// TIA Portal project "DHARMA_1500" (V15) (continued)
VAR_GLOBAL   // PLC tag table "I/O-TurnTable"
   "TT_ES_Operatingpanel" AT %I1104.0 : Bool;   // Turntable: Emergency stop control panel
   "TT_F_CircuitBreaker" AT %I1100.0 : Bool;   // Turntable: Fault supply
   "TT_T_Start" AT %I1104.1 : Bool;   // Turntable: Start automatic
   "TT_T_Stop" AT %I1104.2 : Bool;   // Turntable: Stop automatic
   "TT_T_Reference" AT %I104.5 : Bool;   // Taster zum Turntable: Referezpunktfahren des Rundtisches "Referenzieren"
   "TT_T_TipTT+" AT %I1104.3 : Bool;   // Turntable: Taster Tippen "+" Rundtisch
   "TT_T_TipTT-" AT %I1104.4 : Bool;   // Turntable: Taster Tippen "-" Rundtisch
   "TT_S_OM_Manual" AT %I104.7 : Bool;   // Schlüsselschalter Rundtisch auf Handbetrieb
   "TT_S_OM_Auto" AT %I104.6 : Bool;   // Schlüsselschalter Rundtisch auf Automatikbetrieb
   "TT_B_Empty" AT %I1105.0 : Bool;   // Taster "Leerfahren"
   "TT_B_WithoutFoam" AT %I1105.1 : Bool;   // Taster "ohne schäumen"
   "TT_F_Supply_FC" AT %I1102.4 : Bool;   // Störung der Versorgung des Frequenzumrichters des Rundtisches
   "TT_F_FC" AT %I1101.0 : Bool;   // Turntable: Fault from frequency converter
   "TT_LS_ToolExist" AT %I1102.6 : Bool;   // Lichtschranke Werkzeug bvorhanden
   "TT_LS_ToolClose" AT %I1102.7 : Bool;   // Lichtschranke Werkzeug geschlossen
   "TT_S_SelectDoor_1" AT %I1102.3 : Bool;   // Turntable: Select open door 1
   "TT_AS_WingDoor" AT %I1100.3 : Bool;   // Turntable: Wing dooor rady
   "TT_AS" AT %I1100.7 : Bool;   // Turntable: Automatic stop ready
   "E_MK_Reiniger_Zyl_Aus" AT %I1107.0 : Bool;   // Zylinder 1 Reiniger Mischkopf ausgefahren
   "E_MK_Reiniger_Zyl_Ein" AT %I1107.1 : Bool;   // Zylinder 1 Reiniger Mischkopf eingefahren
   "T_MK_Reiniger_in_GS" AT %I1106.4 : Bool;   // Taster Mischkopfreiniger in Grundstellung fahren
   "T_MK_Reiniger_in_AS" AT %I1106.5 : Bool;   // Taster Mischkopfreiniger in Arbeitsstellung fahren
   "TT_in_position" AT %I1102.5 : Bool;   // Signal "Genauhalt" Rundtisch
   "P_MK_Reiniger_Zyl" AT %I1107.2 : Bool;   // Zylinder 1 Reiniger Mischkopf Druckluft vorhanden
   "TT_Enable_FC" AT %Q104.4 : Bool;   // Ansteuerunr des Umrichters für den Rundtisch
   "TT_V_OpenDoor_1" AT %Q104.2 : Bool;   // Turntable: Clamping valve door 1
   "TT_H_ReleaseDoor_1" AT %Q104.3 : Bool;   // Turntable: Light door 1
   "TT_H_AS" AT %Q105.7 : Bool;   // Turntable: Light automatik stop ready
   "TT_H_Start" AT %Q104.0 : Bool;   // Anzeige zum starten der Anlage
   "TT_H_Anfahrwarnung" AT %Q104.7 : Bool;
   "TT_H_Tip+" AT %Q105.4 : Bool;
   "TT_H_Tip-" AT %Q105.5 : Bool;
   "TT_H_Reference" AT %Q105.6 : Bool;
END_VAR

VAR_GLOBAL   // PLC tag table "I/O TT main"
   "F_fuse_machine(1)" AT %I100.2 : Bool;
   "F_fuse_slip_ring" AT %I100.3 : Bool;
   "ES_turn_table" AT %I100.4 : Bool;
   "AS_turn_table" AT %I100.7 : Bool;
   "F_cooling_unit" AT %I100.5 : Bool;
   "F_fuse_robot" AT %I100.6 : Bool;
   "F_FC_turn_table" AT %I107.0 : Bool;
   "F_fuse_FC_turn_table" AT %I107.1 : Bool;
   "F_fuse_24V_TT_main" AT %I100.1 : Bool;
   "ES_TT_main_cabinet" AT %I101.0 : Bool;
   "ES_TT_operating_panel" AT %I101.1 : Bool;
   "ES_TT_removal_area" AT %I101.2 : Bool;
   "ES_TT_tool_change" AT %I101.3 : Bool;
   "ES_TT_safety_door_robot" AT %I101.4 : Bool;
   "ES_TT_limit_switch_chain" AT %I101.5 : Bool;
   "Controlvoltage_okay" AT %I100.0 : Bool;
   "AS_door_tool_change" AT %I102.0 : Bool;
   "Quit_door_tool_change" AT %I102.1 : Bool;
   "Select_door_tool_change" AT %I102.2 : Bool;
   "AS_door_robot" AT %I102.3 : Bool;
   "Quit_door_robot" AT %I102.4 : Bool;
   "Select_door_robot" AT %I102.5 : Bool;
   "AS_pendelum_flap_to_handling" AT %I102.6 : Bool;
   "AS_pendelum_flap_from_handling" AT %I102.7 : Bool;
   "AS_Scanner_handling" AT %I103.0 : Bool;
   "Button_slider_HP" AT %I103.1 : Bool;
   "Button_slider_WP" AT %I103.2 : Bool;
   "Scanner_dirty" AT %I103.3 : Bool;
   "ES_robot" AT %I101.6 : Bool;
   "AS_robot_safety_area_1" AT %I103.6 : Bool;
   "AS_okay" AT %I103.7 : Bool;
   "ES_foaming_machine" AT %I101.7 : Bool;
   "I_exact_stop_TT" AT %I107.2 : Bool;
   "P_chain_tensioner" AT %I107.3 : Bool;
   "Quit_fault" AT %I104.4 : Bool;
   "Switch_manual_mode" AT %I104.0 : Bool;
   "Switch_automatic_mode" AT %I104.1 : Bool;
   "Button_start_cycle" AT %I104.2 : Bool;
   "Button_stop_cycle" AT %I104.3 : Bool;
   "Button_reference_TT" AT %I105.1 : Bool;
   "Button_TT_empty" AT %I105.2 : Bool;
   "Button_Tip_+" AT %I105.3 : Bool;
   "Button_Tip_-" AT %I105.4 : Bool;
   "Button_extend_cycle" AT %I105.5 : Bool;
   "Button_without_foam" AT %I105.0 : Bool;
   "Button_Move_+" AT %I105.6 : Bool;
   "Button_Move_-" AT %I105.7 : Bool;
   "BCD_Movement_Bit_0" AT %I106.0 : Bool;
   "BCD_Movement_Bit_1" AT %I106.1 : Bool;
   "BCD_Movement_Bit_2" AT %I106.2 : Bool;
   "BCD_Movement_Bit_3" AT %I106.3 : Bool;
   "BCD_MC_Bit_0" AT %I106.4 : Bool;
   "BCD_MC_Bit_1" AT %I106.5 : Bool;
   "BCD_MC_Bit_2" AT %I106.6 : Bool;
   "BCD_MC_Bit_3" AT %I106.7 : Bool;
   "BCD_Movement_MC" AT %IB106 : Byte;
   "Release_FC_turn_table" AT %Q103.7 : Bool;
   "Release_door_tool_change" AT %Q103.0 : Bool;
   "Selected_door_tool_change" AT %Q100.0 : Bool;
   "Release_door_robot" AT %Q103.1 : Bool;
   "Selected_door_robot" AT %Q100.1 : Bool;
   "Quit_scanner_handling" AT %Q100.7 : Bool;
   "LED_slider_HP" AT %Q102.1 : Bool;
   "LED_slider_WP" AT %Q102.2 : Bool;
   "Quit_automatic_stop" AT %Q100.2 : Bool;
   "V_chain_tensioner" AT %Q102.7 : Bool;
   "LED_start_cycle" AT %Q101.0 : Bool;
   "LED_reference_TT" AT %Q101.1 : Bool;
   "LED_TT_empty" AT %Q101.2 : Bool;
   "LED_Tip_+" AT %Q101.3 : Bool;
   "LED_Tip_-" AT %Q101.4 : Bool;
   "LED_extend_cycle" AT %Q101.5 : Bool;
   "LED_Move_+" AT %Q101.6 : Bool;
   "LED_Move_-" AT %Q101.7 : Bool;
   "Horn_TT_start" AT %Q100.3 : Bool;
   "LED_fault" AT %Q100.5 : Bool;
   "Horn_fault" AT %Q100.6 : Bool;
   "LED_TT_ready" AT %Q100.4 : Bool;
END_VAR

VAR_GLOBAL   // PLC tag table "Generell"
   "Flag_10_000_Hertz" AT %M0.0 : Bool;   // System flag of pulse 10.000 Hertz
   "Flag_05_000_Hertz" AT %M0.1 : Bool;   // System flag of pulse 5.000 Hertz
   "Flag_02_500_Hertz" AT %M0.2 : Bool;   // System flag of pulse 2.500 Hertz
   "Flag_02_000_Hertz" AT %M0.3 : Bool;   // System flag of pulse 2.000 Hertz
   "Flag_01_250_Hertz" AT %M0.4 : Bool;   // System flag of pulse 1.250 Hertz
   "Flag_01_000_Hertz" AT %M0.5 : Bool;   // System flag of pulse 1.000 Hertz
   "Flag_00_625_Hertz" AT %M0.6 : Bool;   // System flag of pulse 0.625 Hertz
   "Flag_00_500_Hertz" AT %M0.7 : Bool;   // System flag of pulse 0.500 Hertz
   "Flag_Erster_SPS_Zyklus" AT %M2.1 : Bool;   // Flag first plc cycle running
   "Flag_DP_Bus1_ADR001_ok" AT %M10.0 : Bool;   // profibus member at DP-Bus 01 with address 001 is available
   "Flag_DP_Bus1_ADR002_ok" AT %M10.1 : Bool;   // profibus member at DP-Bus 01 with address 002 is available
   "Flag_DP_Bus1_ADR003_ok" AT %M10.2 : Bool;   // profibus member at DP-Bus 01 with address 003 is available
   "Flag_DP_Bus1_ADR004_ok" AT %M10.3 : Bool;   // profibus member at DP-Bus 01 with address 004 is available
   "Flag_DP_Bus1_ADR005_ok" AT %M10.4 : Bool;   // profibus member at DP-Bus 01 with address 005 is available
   "Flag_DP_Bus1_ADR006_ok" AT %M10.5 : Bool;   // profibus member at DP-Bus 01 with address 006 is available
   "Flag_DP_Bus1_ADR007_ok" AT %M10.6 : Bool;   // profibus member at DP-Bus 01 with address 007 is available
   "Flag_DP_Bus1_ADR008_ok" AT %M10.7 : Bool;   // profibus member at DP-Bus 01 with address 008 is available
   "Flag_DP_Bus1_ADR009_ok" AT %M11.0 : Bool;   // profibus member at DP-Bus 01 with address 009 is available
   "Flag_DP_Bus1_ADR010_ok" AT %M11.1 : Bool;   // profibus member at DP-Bus 01 with address 010 is available
   "Flag_DP_Bus1_ADR011_ok" AT %M11.2 : Bool;   // profibus member at DP-Bus 01 with address 011 is available
   "Flag_DP_Bus1_ADR012_ok" AT %M11.3 : Bool;   // profibus member at DP-Bus 01 with address 012 is available
   "Flag_DP_Bus1_ADR013_ok" AT %M11.4 : Bool;   // profibus member at DP-Bus 01 with address 013 is available
   "Flag_DP_Bus1_ADR014_ok" AT %M11.5 : Bool;   // profibus member at DP-Bus 01 with address 014 is available
   "Flag_DP_Bus1_ADR015_ok" AT %M11.6 : Bool;   // profibus member at DP-Bus 01 with address 015 is available
   "Flag_DP_Bus1_ADR016_ok" AT %M11.7 : Bool;   // profibus member at DP-Bus 01 with address 016 is available
   "Flag_DP_Bus1_ADR017_ok" AT %M12.0 : Bool;   // profibus member at DP-Bus 01 with address 017 is available
   "Flag_DP_Bus1_ADR018_ok" AT %M12.1 : Bool;   // profibus member at DP-Bus 01 with address 018 is available
   "Flag_DP_Bus1_ADR019_ok" AT %M12.2 : Bool;   // profibus member at DP-Bus 01 with address 019 is available
   "Flag_DP_Bus1_ADR020_ok" AT %M12.3 : Bool;   // profibus member at DP-Bus 01 with address 020 is available
   "Flag_DP_Bus1_ADR021_ok" AT %M12.4 : Bool;   // profibus member at DP-Bus 01 with address 021 is available
   "Flag_DP_Bus1_ADR022_ok" AT %M12.5 : Bool;   // profibus member at DP-Bus 01 with address 022 is available
   "Flag_DP_Bus1_ADR023_ok" AT %M12.6 : Bool;   // profibus member at DP-Bus 01 with address 023 is available
   "Flag_DP_Bus1_ADR024_ok" AT %M12.7 : Bool;   // profibus member at DP-Bus 01 with address 024 is available
   "Flag_DP_Bus1_ADR025_ok" AT %M13.0 : Bool;   // profibus member at DP-Bus 01 with address 025 is available
   "Flag_DP_Bus1_ADR026_ok" AT %M13.1 : Bool;   // profibus member at DP-Bus 01 with address 026 is available
   "Flag_DP_Bus1_ADR027_ok" AT %M13.2 : Bool;   // profibus member at DP-Bus 01 with address 027 is available
   "Flag_DP_Bus1_ADR028_ok" AT %M13.3 : Bool;   // profibus member at DP-Bus 01 with address 028 is available
   "Flag_DP_Bus1_ADR029_ok" AT %M13.4 : Bool;   // profibus member at DP-Bus 01 with address 029 is available
   "Flag_DP_Bus1_ADR030_ok" AT %M13.5 : Bool;   // profibus member at DP-Bus 01 with address 030 is available
   "Flag_DP_Bus1_ADR031_ok" AT %M13.6 : Bool;   // profibus member at DP-Bus 01 with address 031 is available
   "Flag_DP_Bus1_ADR032_ok" AT %M13.7 : Bool;   // profibus member at DP-Bus 01 with address 032 is available
   "Flag_DP_Bus1_ADR033_ok" AT %M14.0 : Bool;   // profibus member at DP-Bus 01 with address 033 is available
   "Flag_DP_Bus1_ADR034_ok" AT %M14.1 : Bool;   // profibus member at DP-Bus 01 with address 034 is available
   "Flag_DP_Bus1_ADR035_ok" AT %M14.2 : Bool;   // profibus member at DP-Bus 01 with address 035 is available
   "Flag_DP_Bus1_ADR036_ok" AT %M14.3 : Bool;   // profibus member at DP-Bus 01 with address 036 is available
   "Flag_DP_Bus1_ADR037_ok" AT %M14.4 : Bool;   // profibus member at DP-Bus 01 with address 037 is available
   "Flag_DP_Bus1_ADR038_ok" AT %M14.5 : Bool;   // profibus member at DP-Bus 01 with address 038 is available
   "Flag_DP_Bus1_ADR039_ok" AT %M14.6 : Bool;   // profibus member at DP-Bus 01 with address 039 is available
   "Flag_DP_Bus1_ADR040_ok" AT %M14.7 : Bool;   // profibus member at DP-Bus 01 with address 040 is available
   "Flag_DP_Bus1_ADR041_ok" AT %M15.0 : Bool;   // profibus member at DP-Bus 01 with address 041 is available
   "Flag_DP_Bus1_ADR042_ok" AT %M15.1 : Bool;   // profibus member at DP-Bus 01 with address 042 is available
   "Flag_DP_Bus1_ADR043_ok" AT %M15.2 : Bool;   // profibus member at DP-Bus 01 with address 043 is available
   "Flag_DP_Bus1_ADR044_ok" AT %M15.3 : Bool;   // profibus member at DP-Bus 01 with address 044 is available
   "Flag_DP_Bus1_ADR045_ok" AT %M15.4 : Bool;   // profibus member at DP-Bus 01 with address 045 is available
   "Flag_DP_Bus1_ADR046_ok" AT %M15.5 : Bool;   // profibus member at DP-Bus 01 with address 046 is available
   "Flag_DP_Bus1_ADR047_ok" AT %M15.6 : Bool;   // profibus member at DP-Bus 01 with address 047 is available
   "Flag_DP_Bus1_ADR048_ok" AT %M15.7 : Bool;   // profibus member at DP-Bus 01 with address 048 is available
   "Flag_DP_Bus1_ADR049_ok" AT %M16.0 : Bool;   // profibus member at DP-Bus 01 with address 049 is available
   "Flag_DP_Bus1_ADR050_ok" AT %M16.1 : Bool;   // profibus member at DP-Bus 01 with address 050 is available
   "Flag_DP_Bus1_ADR051_ok" AT %M16.2 : Bool;   // profibus member at DP-Bus 01 with address 051 is available
   "Flag_DP_Bus1_ADR052_ok" AT %M16.3 : Bool;   // profibus member at DP-Bus 01 with address 052 is available
   "Flag_DP_Bus1_ADR053_ok" AT %M16.4 : Bool;   // profibus member at DP-Bus 01 with address 053 is available
   "Flag_DP_Bus1_ADR054_ok" AT %M16.5 : Bool;   // profibus member at DP-Bus 01 with address 054 is available
   "Flag_DP_Bus1_ADR055_ok" AT %M16.6 : Bool;   // profibus member at DP-Bus 01 with address 055 is available
   "Flag_DP_Bus1_ADR056_ok" AT %M16.7 : Bool;   // profibus member at DP-Bus 01 with address 056 is available
   "Flag_DP_Bus1_ADR057_ok" AT %M17.0 : Bool;   // profibus member at DP-Bus 01 with address 057 is available
   "Flag_DP_Bus1_ADR058_ok" AT %M17.1 : Bool;   // profibus member at DP-Bus 01 with address 058 is available
   "Flag_DP_Bus1_ADR059_ok" AT %M17.2 : Bool;   // profibus member at DP-Bus 01 with address 059 is available
   "Flag_DP_Bus1_ADR060_ok" AT %M17.3 : Bool;   // profibus member at DP-Bus 01 with address 060 is available
   "Flag_DP_Bus1_ADR061_ok" AT %M17.4 : Bool;   // profibus member at DP-Bus 01 with address 061 is available
   "Flag_DP_Bus1_ADR062_ok" AT %M17.5 : Bool;   // profibus member at DP-Bus 01 with address 062 is available
   "Flag_DP_Bus1_ADR063_ok" AT %M17.6 : Bool;   // profibus member at DP-Bus 01 with address 063 is available
   "Flag_DP_Bus1_ADR064_ok" AT %M17.7 : Bool;   // profibus member at DP-Bus 01 with address 064 is available
   "Flag_DP_Bus1_ADR065_ok" AT %M18.0 : Bool;   // profibus member at DP-Bus 01 with address 065 is available
   "Flag_DP_Bus1_ADR066_ok" AT %M18.1 : Bool;   // profibus member at DP-Bus 01 with address 066 is available
   "Flag_DP_Bus1_ADR067_ok" AT %M18.2 : Bool;   // profibus member at DP-Bus 01 with address 067 is available
   "Flag_DP_Bus1_ADR068_ok" AT %M18.3 : Bool;   // profibus member at DP-Bus 01 with address 068 is available
   "Flag_DP_Bus1_ADR069_ok" AT %M18.4 : Bool;   // profibus member at DP-Bus 01 with address 069 is available
   "Flag_DP_Bus1_ADR070_ok" AT %M18.5 : Bool;   // profibus member at DP-Bus 01 with address 070 is available
   "Flag_DP_Bus1_ADR071_ok" AT %M18.6 : Bool;   // profibus member at DP-Bus 01 with address 071 is available
   "Flag_DP_Bus1_ADR072_ok" AT %M18.7 : Bool;   // profibus member at DP-Bus 01 with address 072 is available
   "Flag_DP_Bus1_ADR073_ok" AT %M19.0 : Bool;   // profibus member at DP-Bus 01 with address 073 is available
   "Flag_DP_Bus1_ADR074_ok" AT %M19.1 : Bool;   // profibus member at DP-Bus 01 with address 074 is available
   "Flag_DP_Bus1_ADR075_ok" AT %M19.2 : Bool;   // profibus member at DP-Bus 01 with address 075 is available
   "Flag_DP_Bus1_ADR076_ok" AT %M19.3 : Bool;   // profibus member at DP-Bus 01 with address 076 is available
   "Flag_DP_Bus1_ADR077_ok" AT %M19.4 : Bool;   // profibus member at DP-Bus 01 with address 077 is available
   "Flag_DP_Bus1_ADR078_ok" AT %M19.5 : Bool;   // profibus member at DP-Bus 01 with address 078 is available
   "Flag_DP_Bus1_ADR079_ok" AT %M19.6 : Bool;   // profibus member at DP-Bus 01 with address 079 is available
   "Flag_DP_Bus1_ADR080_ok" AT %M19.7 : Bool;   // profibus member at DP-Bus 01 with address 080 is available
   "Flag_DP_Bus1_ADR081_ok" AT %M20.0 : Bool;   // profibus member at DP-Bus 01 with address 081 is available
   "Flag_DP_Bus1_ADR082_ok" AT %M20.1 : Bool;   // profibus member at DP-Bus 01 with address 082 is available
   "Flag_DP_Bus1_ADR083_ok" AT %M20.2 : Bool;   // profibus member at DP-Bus 01 with address 083 is available
   "Flag_DP_Bus1_ADR084_ok" AT %M20.3 : Bool;   // profibus member at DP-Bus 01 with address 084 is available
   "Flag_DP_Bus1_ADR085_ok" AT %M20.4 : Bool;   // profibus member at DP-Bus 01 with address 085 is available
   "Flag_DP_Bus1_ADR086_ok" AT %M20.5 : Bool;   // profibus member at DP-Bus 01 with address 086 is available
   "Flag_DP_Bus1_ADR087_ok" AT %M20.6 : Bool;   // profibus member at DP-Bus 01 with address 087 is available
   "Flag_DP_Bus1_ADR088_ok" AT %M20.7 : Bool;   // profibus member at DP-Bus 01 with address 088 is available
   "Flag_DP_Bus1_ADR089_ok" AT %M21.0 : Bool;   // profibus member at DP-Bus 01 with address 089 is available
   "Flag_DP_Bus1_ADR090_ok" AT %M21.1 : Bool;   // profibus member at DP-Bus 01 with address 090 is available
   "Flag_DP_Bus1_ADR091_ok" AT %M21.2 : Bool;   // profibus member at DP-Bus 01 with address 091 is available
   "Flag_DP_Bus1_ADR092_ok" AT %M21.3 : Bool;   // profibus member at DP-Bus 01 with address 092 is available
   "Flag_DP_Bus1_ADR093_ok" AT %M21.4 : Bool;   // profibus member at DP-Bus 01 with address 093 is available
   "Flag_DP_Bus1_ADR094_ok" AT %M21.5 : Bool;   // profibus member at DP-Bus 01 with address 094 is available
   "Flag_DP_Bus1_ADR095_ok" AT %M21.6 : Bool;   // profibus member at DP-Bus 01 with address 095 is available
   "Flag_DP_Bus1_ADR096_ok" AT %M21.7 : Bool;   // profibus member at DP-Bus 01 with address 096 is available
   "Flag_DP_Bus1_ADR097_ok" AT %M22.0 : Bool;   // profibus member at DP-Bus 01 with address 097 is available
   "Flag_DP_Bus1_ADR098_ok" AT %M22.1 : Bool;   // profibus member at DP-Bus 01 with address 098 is available
   "Flag_DP_Bus1_ADR099_ok" AT %M22.2 : Bool;   // profibus member at DP-Bus 01 with address 099 is available
   "Flag_DP_Bus1_ADR100_ok" AT %M22.3 : Bool;   // profibus member at DP-Bus 01 with address 100 is available
   "Flag_DP_Bus1_ADR101_ok" AT %M22.4 : Bool;   // profibus member at DP-Bus 01 with address 101 is available
   "Flag_DP_Bus1_ADR102_ok" AT %M22.5 : Bool;   // profibus member at DP-Bus 01 with address 102 is available
   "Flag_DP_Bus1_ADR103_ok" AT %M22.6 : Bool;   // profibus member at DP-Bus 01 with address 103 is available
   "Flag_DP_Bus1_ADR104_ok" AT %M22.7 : Bool;   // profibus member at DP-Bus 01 with address 104 is available
   "Flag_DP_Bus1_ADR105_ok" AT %M23.0 : Bool;   // profibus member at DP-Bus 01 with address 105 is available
   "Flag_DP_Bus1_ADR106_ok" AT %M23.1 : Bool;   // profibus member at DP-Bus 01 with address 106 is available
   "Flag_DP_Bus1_ADR107_ok" AT %M23.2 : Bool;   // profibus member at DP-Bus 01 with address 107 is available
   "Flag_DP_Bus1_ADR108_ok" AT %M23.3 : Bool;   // profibus member at DP-Bus 01 with address 108 is available
   "Flag_DP_Bus1_ADR109_ok" AT %M23.4 : Bool;   // profibus member at DP-Bus 01 with address 109 is available
   "Flag_DP_Bus1_ADR110_ok" AT %M23.5 : Bool;   // profibus member at DP-Bus 01 with address 110 is available
   "Flag_DP_Bus1_ADR111_ok" AT %M23.6 : Bool;   // profibus member at DP-Bus 01 with address 111 is available
   "Flag_DP_Bus1_ADR112_ok" AT %M23.7 : Bool;   // profibus member at DP-Bus 01 with address 112 is available
   "Flag_DP_Bus1_ADR113_ok" AT %M24.0 : Bool;   // profibus member at DP-Bus 01 with address 113 is available
   "Flag_DP_Bus1_ADR114_ok" AT %M24.1 : Bool;   // profibus member at DP-Bus 01 with address 114 is available
   "Flag_DP_Bus1_ADR115_ok" AT %M24.2 : Bool;   // profibus member at DP-Bus 01 with address 115 is available
   "Flag_DP_Bus1_ADR116_ok" AT %M24.3 : Bool;   // profibus member at DP-Bus 01 with address 116 is available
   "Flag_DP_Bus1_ADR117_ok" AT %M24.4 : Bool;   // profibus member at DP-Bus 01 with address 117 is available
   "Flag_DP_Bus1_ADR118_ok" AT %M24.5 : Bool;   // profibus member at DP-Bus 01 with address 118 is available
   "Flag_DP_Bus1_ADR119_ok" AT %M24.6 : Bool;   // profibus member at DP-Bus 01 with address 119 is available
   "Flag_DP_Bus1_ADR120_ok" AT %M24.7 : Bool;   // profibus member at DP-Bus 01 with address 120 is available
   "Flag_DP_Bus1_ADR121_ok" AT %M25.0 : Bool;   // profibus member at DP-Bus 01 with address 121 is available
   "Flag_DP_Bus1_ADR122_ok" AT %M25.1 : Bool;   // profibus member at DP-Bus 01 with address 122 is available
   "Flag_DP_Bus1_ADR123_ok" AT %M25.2 : Bool;   // profibus member at DP-Bus 01 with address 123 is available
   "Flag_DP_Bus1_ADR124_ok" AT %M25.3 : Bool;   // profibus member at DP-Bus 01 with address 124 is available
   "Flag_DP_Bus1_ADR125_ok" AT %M25.4 : Bool;   // profibus member at DP-Bus 01 with address 125 is available
   "Flag_DP_Bus1_ADR126_ok" AT %M25.5 : Bool;   // profibus member at DP-Bus 01 with address 126 is available
   "Flag_DP_Bus1_ADR127_ok" AT %M25.6 : Bool;   // profibus member at DP-Bus 01 with address 127 is available
   "Flag_DP_Bus1_ADR128_ok" AT %M25.7 : Bool;   // profibus member at DP-Bus 01 with address 128 is available
   "Clock_Byte" AT %MB0 : Byte;
   "System_Byte" AT %MB1 : Byte;
   "FirstScan" AT %M1.0 : Bool;
   "DiagStatusUpdate" AT %M1.1 : Bool;
   "AlwaysTRUE" AT %M1.2 : Bool;
   "AlwaysFALSE" AT %M1.3 : Bool;
END_VAR

VAR_GLOBAL   // PLC tag table "Maschinenbett K1/2"
   "M_RTM0Running" AT %M2.0 : Bool;
   "HF_FP_SwitchOffPump" AT %M110.4 : Bool;
   "PulsePumpSwitchedOff" AT %M110.3 : Bool;
   "ShotDisabledDuringShot" AT %M190.0 : Bool;
   "HF_ShotDisabledDuringShot" AT %M190.1 : Bool;
   "HF_FP_ShotRunning" AT %M190.2 : Bool;
   "H_Ready_for_Operation_M1" AT %M90.0 : Bool;
   "H_Ready_for_Operation_M2" AT %M90.1 : Bool;
END_VAR

VAR_GLOBAL   // PLC tag table "E/A- Belegung PW"
   "C_DayTank_C2" AT %IW512 : Int;
   "C_DayTank_C1" AT %IW514 : Int;
   "P_Pump_C1" AT %IW520 : Int;
   "P_Pump_C2" AT %IW522 : Int;
   "L_DayTank_C1" AT %IW524 : Int;
   "L_DayTank_C2" AT %IW526 : Int;
   "C_HeatExchange_C1" AT %IW516 : Int;
   "C_HeatExchange_C2" AT %IW518 : Int;
   "F_air" AT %IW330 : Int;   // Inlet flow air
   "Set_FeedingP_C1" AT %QW516 : Int;
   "Set_FeedingP_C2" AT %QW518 : Int;
END_VAR

VAR_GLOBAL   // PLC tag table "FRA_Int"
   "Interface_Signals_From_KMI" AT %IW100 : Word;
   "FRA_KM_input" AT %I700.0 : "UDT2001_Input_Faurecia";
   "Alarm_Bits_to_KMI" AT %QW230 : Word;
   "Interface_Signals_TO_KMI" AT %QW240 : Word;
   "MH_Number_to_KMI" AT %QW200 : Word;
   "Shotwight_to_KMI" AT %QW202 : Word;
   "Shottime_to_KMI" AT %QW204 : Word;
   "Temp_C1_MH_to_KMI" AT %QW206 : Word;
   "Temp_C2_MH_to_KMI" AT %QW208 : Word;
   "Ratio_C1_to_KMI" AT %QW214 : Word;
   "Ratio_C2_to_KMI" AT %QW216 : Word;
   "Pressure_C1_MH_to_KMI" AT %QW222 : Word;
   "Pressure_C2_MH_to_KMI" AT %QW224 : Word;
   "FRA_KM_output" AT %Q700.0 : "UDT2002_Output_Faurecia";
   "Exp_Ok" AT %MW111 : Int;
   "CP_forward" AT %MW114 : Int;
   "CP_is_forward" AT %MW116 : Int;
   "cycle_run" AT %MW118 : Int;
   "MH_open" AT %MW126 : Int;
   "MHAutomatic" AT %MW128 : Int;
   "Preperation" AT %MW130 : Int;
   "PU_Ok" AT %MW132 : Int;
   "ReadyForShot" AT %MW136 : Int;
   "ServiceMode" AT %MW140 : Int;
   "ShotEnd" AT %MW142 : Int;
   "ShotRun" AT %MW144 : Int;
   "Stop" AT %MW150 : Int;
   "Strobe" AT %MW152 : Int;
   "StrobeQuitt" AT %MW154 : Int;
   "StrobeInv" AT %MW156 : Int;
   "Helpflag_Send_Data_KMI" AT %M166.0 : Bool;
   "Send_Data_to_KMI" AT %M166.1 : Bool;
   "FRA_KM_HM_FP_Circulation" AT %M100.1 : Bool;   // Hilfsmerker positive Flanke reduzierter Betrieb von der Schnittstelle
   "FRA_KM_Quitt" AT %M100.0 : Bool;
   "FRA_KM_HM_FP_Betrieb" AT %M82.2 : Bool;   // Hilfsmerker positive Flanke Service Betrieb von der Schnittstelle
   "FRA_KM_HM_FP_STROBE" AT %M100.2 : Bool;   // Hilfsmerker positive Flanke Start von der Schnittstelle
   "FRA_KM_FP_STROBE" AT %M100.3 : Bool;   // positive Flanke Start von der Schnittstelle
   "FRA_KM_STG_Data" AT %M100.4 : Bool;   // Störung Daten einlöesen
   "FRA_KM_FP_Circulation" AT %M100.5 : Bool;   // positive Flanke reduzierter Betrieb von der Schnittstelle
   "FRA_KM_FP_Betrieb" AT %M82.3 : Bool;   // positive Flanke Service Betrieb von der Schnittstelle
END_VAR
